(* Logix 5000 project; controller MV vendor 1 type 14 code 217 rev 31.11; software revision 31.00; part 31 of 53 *)
(* tags used below, declared in another part *)
   Alarm_Reset : BOOL;
   CWD : CHECKWORD_FLAGS;
   Default_Check_Time : DINT;
   Item_Faults_Are_Latched : BOOL;
   Item_Simulation_Flag : BOOL;
   MC_CD_T1 : PlantItem;   // CD_T1
   MC_CD_T1_ALARM : ALARM_DIGITAL;
   MC_CD_T1_C : ALIAS FOR RIO_Rack_2:7:I.Data.23;
   MC_CD_T1_DR : ALIAS FOR RIO_Rack_2:8:O.Data.11;
   MC_CD_T1_O : ALIAS FOR RIO_Rack_2:7:I.Data.19;
   MC_CD_T2 : PlantItem;   // CD_T2
   MC_CD_T2_ALARM : ALARM_DIGITAL;
   MC_CD_T2_C : ALIAS FOR RIO_Rack_2:7:I.Data.28;
   MC_CD_T2_DR : ALIAS FOR RIO_Rack_2:8:O.Data.12;
   MC_CD_T2_O : ALIAS FOR RIO_Rack_2:7:I.Data.24;
   MC_CH2_DR1 : PlantItem;   // CH2_DR1
   MC_CH2_DR1_ALARM : ALARM_DIGITAL;
   MC_CH2_DR1_C : ALIAS FOR RIO_Rack_2:7:I.Data.6;
   MC_CH2_DR1_DR : ALIAS FOR RIO_Rack_2:8:O.Data.2;
   MC_CH2_DR1_O : ALIAS FOR RIO_Rack_2:7:I.Data.2;
   MC_CH2_DR2 : PlantItem;   // CH2_DR2
   MC_CH2_DR2_ALARM : ALARM_DIGITAL;
   MC_CH2_DR2_C : ALIAS FOR RIO_Rack_2:7:I.Data.7;
   MC_CH2_DR2_DR : ALIAS FOR RIO_Rack_2:8:O.Data.3;
   MC_CH2_DR2_O : ALIAS FOR RIO_Rack_2:7:I.Data.3;
   MC_CH2_DRAIN : PlantItem;   // CH2_DRAIN
   MC_CH2_DRAIN_ALARM : ALARM_DIGITAL;
   MC_CH2_DRAIN_C : ALIAS FOR RIO_Rack_2:7:I.Data.4;
   MC_CH2_DRAIN_DR : ALIAS FOR RIO_Rack_2:8:O.Data.0;
   MC_CH2_DRAIN_O : ALIAS FOR RIO_Rack_2:7:I.Data.0;
   MC_CH2_DT1 : PlantItem;   // CH2_DT1
   MC_CH2_DT1_ALARM : ALARM_DIGITAL;
   MC_CH2_DT1_C : ALIAS FOR RIO_Rack_2:7:I.Data.12;
   MC_CH2_DT1_DR : ALIAS FOR RIO_Rack_2:8:O.Data.4;
   MC_CH2_DT1_O : ALIAS FOR RIO_Rack_2:7:I.Data.8;
   MC_CH2_DT2 : PlantItem;   // CH2_DT2
   MC_CH2_DT2_ALARM : ALARM_DIGITAL;
   MC_CH2_DT2_C : ALIAS FOR RIO_Rack_2:7:I.Data.13;
   MC_CH2_DT2_DR : ALIAS FOR RIO_Rack_2:8:O.Data.5;
   MC_CH2_DT2_O : ALIAS FOR RIO_Rack_2:7:I.Data.9;
   MC_CH2_LF1 : PlantItem;   // CH2_LF1
   MC_CH2_LF1_ALARM : ALARM_DIGITAL;
   MC_CH2_LF1_C : ALIAS FOR RIO_Rack_2:7:I.Data.15;
   MC_CH2_LF1_DR : ALIAS FOR RIO_Rack_2:8:O.Data.7;
   MC_CH2_LF1_O : ALIAS FOR RIO_Rack_2:7:I.Data.11;
   MC_CH2_PR1 : PlantItem;   // CH2_PR1
   MC_CH2_PR1_ALARM : ALARM_DIGITAL;
   MC_CH2_PR1_C : ALIAS FOR RIO_Rack_2:7:I.Data.14;
   MC_CH2_PR1_DR : ALIAS FOR RIO_Rack_2:8:O.Data.6;
   MC_CH2_PR1_O : ALIAS FOR RIO_Rack_2:7:I.Data.10;
   MC_CH2_R6R : PlantItem;   // CH2_R6R
   MC_CH2_R6R_ALARM : ALARM_DIGITAL;
   MC_CH2_R6R_C : ALIAS FOR RIO_Rack_2:6:I.Data.31;
   MC_CH2_R6R_DR : ALIAS FOR RIO_Rack_2:5:O.Data.31;
   MC_CH2_R6R_O : ALIAS FOR RIO_Rack_2:6:I.Data.27;
   MC_CH2_RR : PlantItem;   // CH2_RR
   MC_CH2_RR_ALARM : ALARM_DIGITAL;
   MC_CH2_RR_C : ALIAS FOR RIO_Rack_2:7:I.Data.5;
   MC_CH2_RR_DR : ALIAS FOR RIO_Rack_2:8:O.Data.1;
   MC_CH2_RR_O : ALIAS FOR RIO_Rack_2:7:I.Data.1;
   MC_FL_D1 : PlantItem;   // FL_D1
   MC_FL_D1_ALARM : ALARM_DIGITAL;
   MC_FL_D1_C : ALIAS FOR RIO_Rack_2:7:I.Data.21;
   MC_FL_D1_DR : ALIAS FOR RIO_Rack_2:8:O.Data.9;
   MC_FL_D1_O : ALIAS FOR RIO_Rack_2:7:I.Data.17;
   MC_FL_D2 : PlantItem;   // FL_D2
   MC_FL_D2_ALARM : ALARM_DIGITAL;
   MC_FL_D2_C : ALIAS FOR RIO_Rack_2:7:I.Data.22;
   MC_FL_D2_DR : ALIAS FOR RIO_Rack_2:8:O.Data.10;
   MC_FL_D2_O : ALIAS FOR RIO_Rack_2:7:I.Data.18;
   MC_FL_PR : PlantItem;   // FL_PR
   MC_FL_PR_ALARM : ALARM_DIGITAL;
   MC_FL_PR_C : ALIAS FOR RIO_Rack_2:7:I.Data.20;
   MC_FL_PR_DR : ALIAS FOR RIO_Rack_2:8:O.Data.8;
   MC_FL_PR_O : ALIAS FOR RIO_Rack_2:7:I.Data.16;
   MC_R3S_DR : PlantItem;   // R3S_DR
   MC_R3S_DR_ALARM : ALARM_DIGITAL;
   MC_R3S_DR_C : ALIAS FOR RIO_Rack_2:9:I.Data.15;
   MC_R3S_DR_DR : ALIAS FOR RIO_Rack_2:8:O.Data.23;
   MC_R3S_DR_O : ALIAS FOR RIO_Rack_2:9:I.Data.11;
   MC_R3V1 : PlantItem;   // R3V1
   MC_R3V1_ALARM : ALARM_DIGITAL;
   MC_R3V1_C : ALIAS FOR RIO_Rack_2:9:I.Data.12;
   MC_R3V1_DR : ALIAS FOR RIO_Rack_2:8:O.Data.20;
   MC_R3V1_O : ALIAS FOR RIO_Rack_2:9:I.Data.8;
   MC_R3V2 : PlantItem;   // R3V2
   MC_R3V2_ALARM : ALARM_DIGITAL;
   MC_R3V2_C : ALIAS FOR RIO_Rack_2:9:I.Data.13;
   MC_R3V2_DR : ALIAS FOR RIO_Rack_2:8:O.Data.21;
   MC_R3V2_O : ALIAS FOR RIO_Rack_2:9:I.Data.9;
   MC_SPV1 : PlantItem;   // SPV1
   MC_SPV1_ALARM : ALARM_DIGITAL;
   MC_SPV1_C : ALIAS FOR RIO_Rack_2:7:I.Data.31;
   MC_SPV1_DR : ALIAS FOR RIO_Rack_2:8:O.Data.15;
   MC_SPV1_O : ALIAS FOR RIO_Rack_2:7:I.Data.27;
   MC_SPV2 : PlantItem;   // SPV2
   MC_SPV2_ALARM : ALARM_DIGITAL;
   MC_SPV2_C : ALIAS FOR RIO_Rack_2:9:I.Data.4;
   MC_SPV2_DR : ALIAS FOR RIO_Rack_2:8:O.Data.16;
   MC_SPV2_O : ALIAS FOR RIO_Rack_2:9:I.Data.0;
   MC_SPV3 : PlantItem;   // SPV3
   MC_SPV3_ALARM : ALARM_DIGITAL;
   MC_SPV3_C : ALIAS FOR RIO_Rack_2:9:I.Data.5;
   MC_SPV3_DR : ALIAS FOR RIO_Rack_2:8:O.Data.17;
   MC_SPV3_O : ALIAS FOR RIO_Rack_2:9:I.Data.1;
   MC_SPV4 : PlantItem;   // SPV4
   MC_SPV4_ALARM : ALARM_DIGITAL;
   MC_SPV4_C : ALIAS FOR RIO_Rack_2:9:I.Data.6;
   MC_SPV4_DR : ALIAS FOR RIO_Rack_2:8:O.Data.18;
   MC_SPV4_O : ALIAS FOR RIO_Rack_2:9:I.Data.2;
   MC_SPV5 : PlantItem;   // SPV5
   MC_SPV5_ALARM : ALARM_DIGITAL;
   MC_SPV5_C : ALIAS FOR RIO_Rack_2:9:I.Data.7;
   MC_SPV5_DR : ALIAS FOR RIO_Rack_2:8:O.Data.19;
   MC_SPV5_O : ALIAS FOR RIO_Rack_2:9:I.Data.3;
   MC_SV1 : PlantItem;   // SV1
   MC_SV1_ALARM : ALARM_DIGITAL;
   MC_SV1_C : ALIAS FOR RIO_Rack_2:7:I.Data.29;
   MC_SV1_DR : ALIAS FOR RIO_Rack_2:8:O.Data.13;
   MC_SV1_O : ALIAS FOR RIO_Rack_2:7:I.Data.25;
   MC_SV2 : PlantItem;   // SV2
   MC_SV2_ALARM : ALARM_DIGITAL;
   MC_SV2_C : ALIAS FOR RIO_Rack_2:7:I.Data.30;
   MC_SV2_DR : ALIAS FOR RIO_Rack_2:8:O.Data.14;
   MC_SV2_O : ALIAS FOR RIO_Rack_2:7:I.Data.26;
   One_Second_One_Scan : ALIAS FOR One_Second_1_scan;
(* MC_Common, continued *)

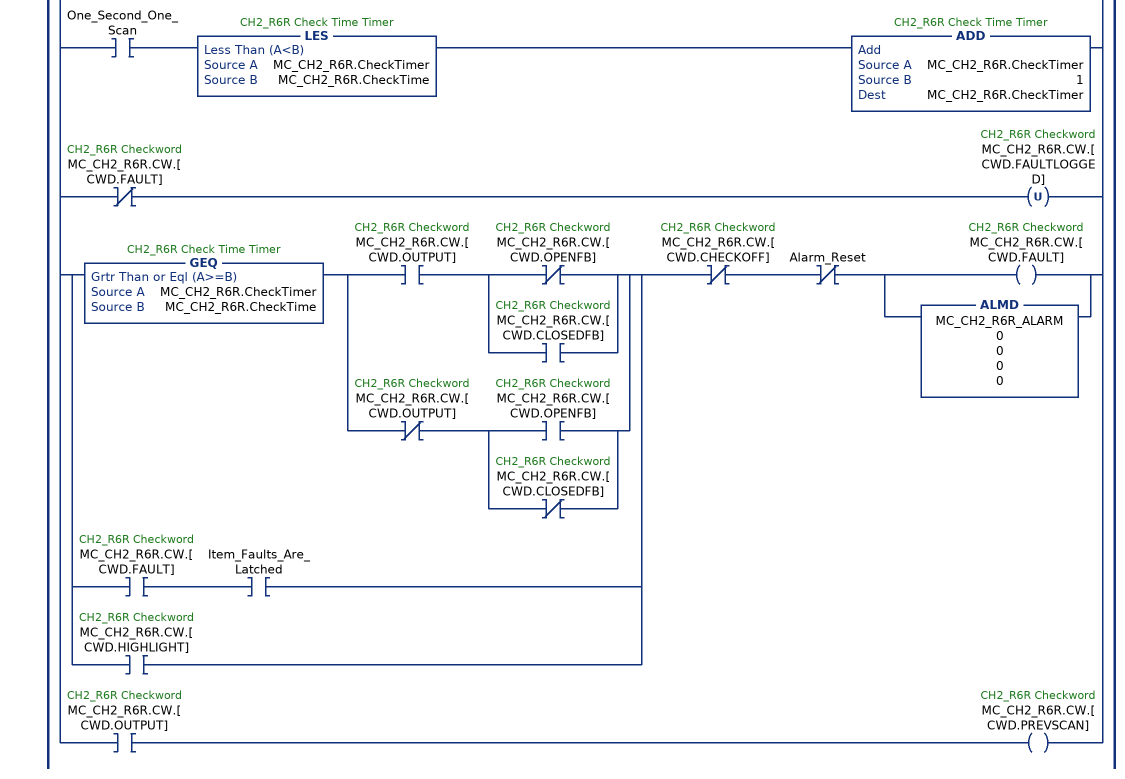
   [picture p660: MC_Common/MC_Valves rungs 31-31]
   31: [NEQ(MC_CH2_R6R.DriveBits,0) OTE(MC_CH2_R6R.CW.[CWD.AUTODRV]) ,[XIC(MC_CH2_R6R.CW.[CWD.AUTODRV]) XIO(MC_CH2_R6R.CW.[CWD.MANUAL]) ,XIC(MC_CH2_R6R.CW.[CWD.MANDRV]) XIC(MC_CH2_R6R.CW.[CWD.MANUAL]) ] OTE(MC_CH2_R6R.CW.[CWD.OUTPUT]) ,XIC(MC_CH2_R6R.CW.[CWD.OUTPUT]) OTE(MC_CH2_R6R_DR) ,XIC(S:FS) [OTU(MC_CH2_R6R.CW.[CWD.MANUAL]) ,LEQ(MC_CH2_R6R.CheckTime,0) MOV(Default_Check_Time,MC_CH2_R6R.CheckTime) ] ,[[XIC(MC_CH2_R6R_O) XIO(Item_Simulation_Flag) ,XIC(Item_Simulation_Flag) XIC(MC_CH2_R6R.CW.[CWD.OUTPUT]) XIO(MC_CH2_R6R.CW.[CWD.SIMFAIL]) ] OTE(MC_CH2_R6R.CW.[CWD.OPENFB]) ,[XIC(MC_CH2_R6R_C) XIO(Item_Simulation_Flag) ,XIC(Item_Simulation_Flag) XIO(MC_CH2_R6R.CW.[CWD.OUTPUT]) XIO(MC_CH2_R6R.CW.[CWD.SIMFAIL]) ] OTE(MC_CH2_R6R.CW.[CWD.CLOSEDFB]) ] ,[XIC(MC_CH2_R6R.CW.[CWD.OUTPUT]) XIO(MC_CH2_R6R.CW.[CWD.PREVSCAN]) ,XIO(MC_CH2_R6R.CW.[CWD.OUTPUT]) XIC(MC_CH2_R6R.CW.[CWD.PREVSCAN]) ] CLR(MC_CH2_R6R.CheckTimer) ,XIC(One_Second_One_Scan) LES(MC_CH2_R6R.CheckTimer,MC_CH2_R6R.CheckTime) ADD(MC_CH2_R6R.CheckTimer,1,MC_CH2_R6R.CheckTimer) ,XIO(MC_CH2_R6R.CW.[CWD.FAULT]) OTU(MC_CH2_R6R.CW.[CWD.FAULTLOGGED]) ,[GEQ(MC_CH2_R6R.CheckTimer,MC_CH2_R6R.CheckTime) [XIC(MC_CH2_R6R.CW.[CWD.OUTPUT]) [XIO(MC_CH2_R6R.CW.[CWD.OPENFB]) ,XIC(MC_CH2_R6R.CW.[CWD.CLOSEDFB]) ] ,XIO(MC_CH2_R6R.CW.[CWD.OUTPUT]) [XIC(MC_CH2_R6R.CW.[CWD.OPENFB]) ,XIO(MC_CH2_R6R.CW.[CWD.CLOSEDFB]) ] ] ,XIC(MC_CH2_R6R.CW.[CWD.FAULT]) XIC(Item_Faults_Are_Latched) ,XIC(MC_CH2_R6R.CW.[CWD.HIGHLIGHT]) ] XIO(MC_CH2_R6R.CW.[CWD.CHECKOFF]) XIO(Alarm_Reset) [OTE(MC_CH2_R6R.CW.[CWD.FAULT]) ,ALMD(MC_CH2_R6R_ALARM,0,0,0,0) ] ,XIC(MC_CH2_R6R.CW.[CWD.OUTPUT]) OTE(MC_CH2_R6R.CW.[CWD.PREVSCAN]) ];
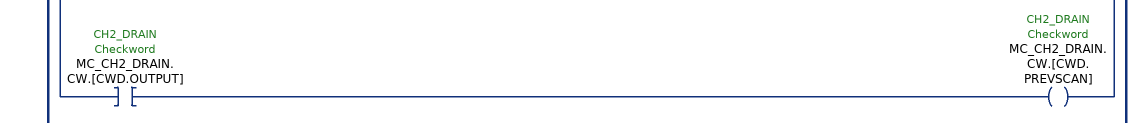
   32: [NEQ(MC_CH2_DRAIN.DriveBits,0) OTE(MC_CH2_DRAIN.CW.[CWD.AUTODRV]) ,[XIC(MC_CH2_DRAIN.CW.[CWD.AUTODRV]) XIO(MC_CH2_DRAIN.CW.[CWD.MANUAL]) ,XIC(MC_CH2_DRAIN.CW.[CWD.MANDRV]) XIC(MC_CH2_DRAIN.CW.[CWD.MANUAL]) ] OTE(MC_CH2_DRAIN.CW.[CWD.OUTPUT]) ,XIC(MC_CH2_DRAIN.CW.[CWD.OUTPUT]) OTE(MC_CH2_DRAIN_DR) ,XIC(S:FS) [OTU(MC_CH2_DRAIN.CW.[CWD.MANUAL]) ,LEQ(MC_CH2_DRAIN.CheckTime,0) MOV(Default_Check_Time,MC_CH2_DRAIN.CheckTime) ] ,[[XIC(MC_CH2_DRAIN_O) XIO(Item_Simulation_Flag) ,XIC(Item_Simulation_Flag) XIC(MC_CH2_DRAIN.CW.[CWD.OUTPUT]) XIO(MC_CH2_DRAIN.CW.[CWD.SIMFAIL]) ] OTE(MC_CH2_DRAIN.CW.[CWD.OPENFB]) ,[XIC(MC_CH2_DRAIN_C) XIO(Item_Simulation_Flag) ,XIC(Item_Simulation_Flag) XIO(MC_CH2_DRAIN.CW.[CWD.OUTPUT]) XIO(MC_CH2_DRAIN.CW.[CWD.SIMFAIL]) ] OTE(MC_CH2_DRAIN.CW.[CWD.CLOSEDFB]) ] ,[XIC(MC_CH2_DRAIN.CW.[CWD.OUTPUT]) XIO(MC_CH2_DRAIN.CW.[CWD.PREVSCAN]) ,XIO(MC_CH2_DRAIN.CW.[CWD.OUTPUT]) XIC(MC_CH2_DRAIN.CW.[CWD.PREVSCAN]) ] CLR(MC_CH2_DRAIN.CheckTimer) ,XIC(One_Second_One_Scan) LES(MC_CH2_DRAIN.CheckTimer,MC_CH2_DRAIN.CheckTime) ADD(MC_CH2_DRAIN.CheckTimer,1,MC_CH2_DRAIN.CheckTimer) ,XIO(MC_CH2_DRAIN.CW.[CWD.FAULT]) OTU(MC_CH2_DRAIN.CW.[CWD.FAULTLOGGED]) ,[GEQ(MC_CH2_DRAIN.CheckTimer,MC_CH2_DRAIN.CheckTime) [XIC(MC_CH2_DRAIN.CW.[CWD.OUTPUT]) [XIO(MC_CH2_DRAIN.CW.[CWD.OPENFB]) ,XIC(MC_CH2_DRAIN.CW.[CWD.CLOSEDFB]) ] ,XIO(MC_CH2_DRAIN.CW.[CWD.OUTPUT]) [XIC(MC_CH2_DRAIN.CW.[CWD.OPENFB]) ,XIO(MC_CH2_DRAIN.CW.[CWD.CLOSEDFB]) ] ] ,XIC(MC_CH2_DRAIN.CW.[CWD.FAULT]) XIC(Item_Faults_Are_Latched) ,XIC(MC_CH2_DRAIN.CW.[CWD.HIGHLIGHT]) ] XIO(MC_CH2_DRAIN.CW.[CWD.CHECKOFF]) XIO(Alarm_Reset) [OTE(MC_CH2_DRAIN.CW.[CWD.FAULT]) ,ALMD(MC_CH2_DRAIN_ALARM,0,0,0,0) ] ,XIC(MC_CH2_DRAIN.CW.[CWD.OUTPUT]) OTE(MC_CH2_DRAIN.CW.[CWD.PREVSCAN]) ];
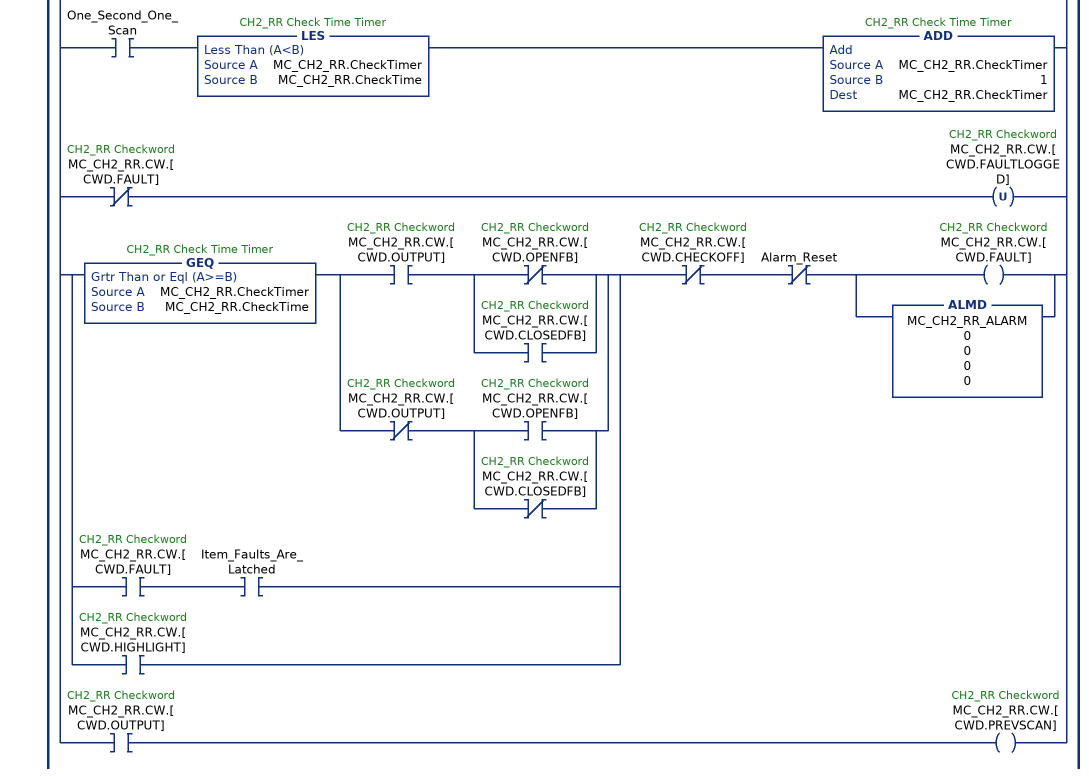
   33: [NEQ(MC_CH2_RR.DriveBits,0) OTE(MC_CH2_RR.CW.[CWD.AUTODRV]) ,[XIC(MC_CH2_RR.CW.[CWD.AUTODRV]) XIO(MC_CH2_RR.CW.[CWD.MANUAL]) ,XIC(MC_CH2_RR.CW.[CWD.MANDRV]) XIC(MC_CH2_RR.CW.[CWD.MANUAL]) ] OTE(MC_CH2_RR.CW.[CWD.OUTPUT]) ,XIC(MC_CH2_RR.CW.[CWD.OUTPUT]) OTE(MC_CH2_RR_DR) ,XIC(S:FS) [OTU(MC_CH2_RR.CW.[CWD.MANUAL]) ,LEQ(MC_CH2_RR.CheckTime,0) MOV(Default_Check_Time,MC_CH2_RR.CheckTime) ] ,[[XIC(MC_CH2_RR_O) XIO(Item_Simulation_Flag) ,XIC(Item_Simulation_Flag) XIC(MC_CH2_RR.CW.[CWD.OUTPUT]) XIO(MC_CH2_RR.CW.[CWD.SIMFAIL]) ] OTE(MC_CH2_RR.CW.[CWD.OPENFB]) ,[XIC(MC_CH2_RR_C) XIO(Item_Simulation_Flag) ,XIC(Item_Simulation_Flag) XIO(MC_CH2_RR.CW.[CWD.OUTPUT]) XIO(MC_CH2_RR.CW.[CWD.SIMFAIL]) ] OTE(MC_CH2_RR.CW.[CWD.CLOSEDFB]) ] ,[XIC(MC_CH2_RR.CW.[CWD.OUTPUT]) XIO(MC_CH2_RR.CW.[CWD.PREVSCAN]) ,XIO(MC_CH2_RR.CW.[CWD.OUTPUT]) XIC(MC_CH2_RR.CW.[CWD.PREVSCAN]) ] CLR(MC_CH2_RR.CheckTimer) ,XIC(One_Second_One_Scan) LES(MC_CH2_RR.CheckTimer,MC_CH2_RR.CheckTime) ADD(MC_CH2_RR.CheckTimer,1,MC_CH2_RR.CheckTimer) ,XIO(MC_CH2_RR.CW.[CWD.FAULT]) OTU(MC_CH2_RR.CW.[CWD.FAULTLOGGED]) ,[GEQ(MC_CH2_RR.CheckTimer,MC_CH2_RR.CheckTime) [XIC(MC_CH2_RR.CW.[CWD.OUTPUT]) [XIO(MC_CH2_RR.CW.[CWD.OPENFB]) ,XIC(MC_CH2_RR.CW.[CWD.CLOSEDFB]) ] ,XIO(MC_CH2_RR.CW.[CWD.OUTPUT]) [XIC(MC_CH2_RR.CW.[CWD.OPENFB]) ,XIO(MC_CH2_RR.CW.[CWD.CLOSEDFB]) ] ] ,XIC(MC_CH2_RR.CW.[CWD.FAULT]) XIC(Item_Faults_Are_Latched) ,XIC(MC_CH2_RR.CW.[CWD.HIGHLIGHT]) ] XIO(MC_CH2_RR.CW.[CWD.CHECKOFF]) XIO(Alarm_Reset) [OTE(MC_CH2_RR.CW.[CWD.FAULT]) ,ALMD(MC_CH2_RR_ALARM,0,0,0,0) ] ,XIC(MC_CH2_RR.CW.[CWD.OUTPUT]) OTE(MC_CH2_RR.CW.[CWD.PREVSCAN]) ];
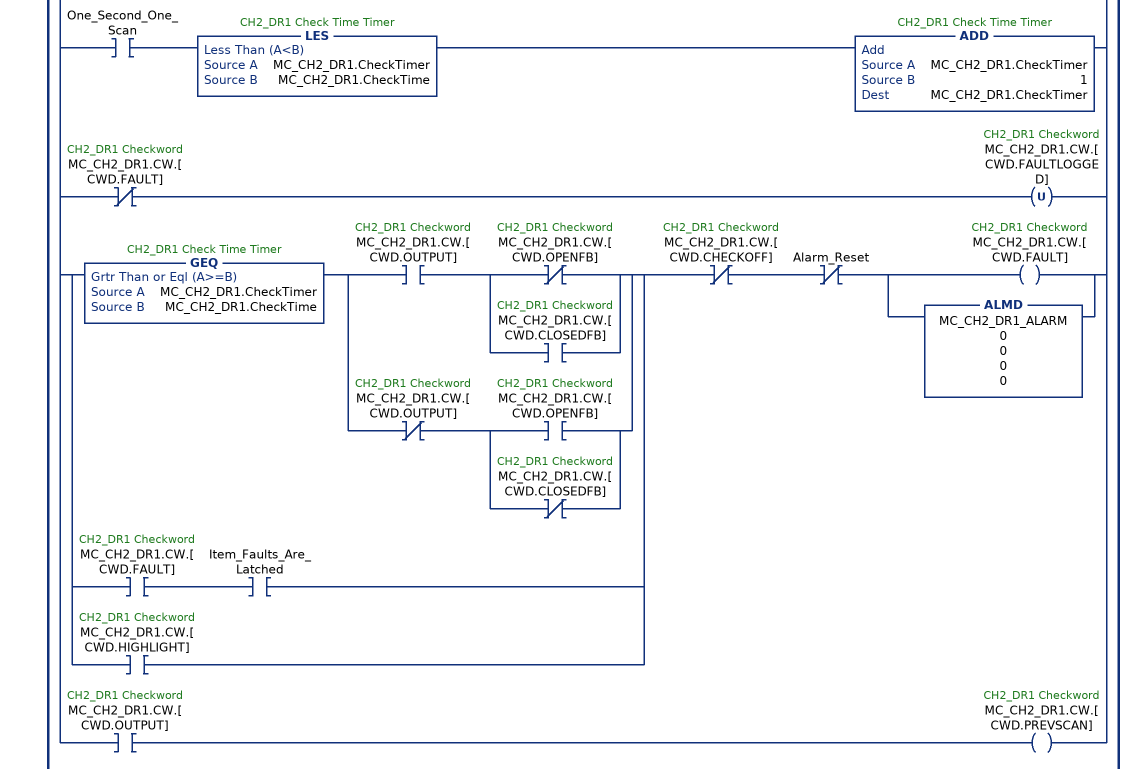
   34: [NEQ(MC_CH2_DR1.DriveBits,0) OTE(MC_CH2_DR1.CW.[CWD.AUTODRV]) ,[XIC(MC_CH2_DR1.CW.[CWD.AUTODRV]) XIO(MC_CH2_DR1.CW.[CWD.MANUAL]) ,XIC(MC_CH2_DR1.CW.[CWD.MANDRV]) XIC(MC_CH2_DR1.CW.[CWD.MANUAL]) ] OTE(MC_CH2_DR1.CW.[CWD.OUTPUT]) ,XIC(MC_CH2_DR1.CW.[CWD.OUTPUT]) OTE(MC_CH2_DR1_DR) ,XIC(S:FS) [OTU(MC_CH2_DR1.CW.[CWD.MANUAL]) ,LEQ(MC_CH2_DR1.CheckTime,0) MOV(Default_Check_Time,MC_CH2_DR1.CheckTime) ] ,[[XIC(MC_CH2_DR1_O) XIO(Item_Simulation_Flag) ,XIC(Item_Simulation_Flag) XIC(MC_CH2_DR1.CW.[CWD.OUTPUT]) XIO(MC_CH2_DR1.CW.[CWD.SIMFAIL]) ] OTE(MC_CH2_DR1.CW.[CWD.OPENFB]) ,[XIC(MC_CH2_DR1_C) XIO(Item_Simulation_Flag) ,XIC(Item_Simulation_Flag) XIO(MC_CH2_DR1.CW.[CWD.OUTPUT]) XIO(MC_CH2_DR1.CW.[CWD.SIMFAIL]) ] OTE(MC_CH2_DR1.CW.[CWD.CLOSEDFB]) ] ,[XIC(MC_CH2_DR1.CW.[CWD.OUTPUT]) XIO(MC_CH2_DR1.CW.[CWD.PREVSCAN]) ,XIO(MC_CH2_DR1.CW.[CWD.OUTPUT]) XIC(MC_CH2_DR1.CW.[CWD.PREVSCAN]) ] CLR(MC_CH2_DR1.CheckTimer) ,XIC(One_Second_One_Scan) LES(MC_CH2_DR1.CheckTimer,MC_CH2_DR1.CheckTime) ADD(MC_CH2_DR1.CheckTimer,1,MC_CH2_DR1.CheckTimer) ,XIO(MC_CH2_DR1.CW.[CWD.FAULT]) OTU(MC_CH2_DR1.CW.[CWD.FAULTLOGGED]) ,[GEQ(MC_CH2_DR1.CheckTimer,MC_CH2_DR1.CheckTime) [XIC(MC_CH2_DR1.CW.[CWD.OUTPUT]) [XIO(MC_CH2_DR1.CW.[CWD.OPENFB]) ,XIC(MC_CH2_DR1.CW.[CWD.CLOSEDFB]) ] ,XIO(MC_CH2_DR1.CW.[CWD.OUTPUT]) [XIC(MC_CH2_DR1.CW.[CWD.OPENFB]) ,XIO(MC_CH2_DR1.CW.[CWD.CLOSEDFB]) ] ] ,XIC(MC_CH2_DR1.CW.[CWD.FAULT]) XIC(Item_Faults_Are_Latched) ,XIC(MC_CH2_DR1.CW.[CWD.HIGHLIGHT]) ] XIO(MC_CH2_DR1.CW.[CWD.CHECKOFF]) XIO(Alarm_Reset) [OTE(MC_CH2_DR1.CW.[CWD.FAULT]) ,ALMD(MC_CH2_DR1_ALARM,0,0,0,0) ] ,XIC(MC_CH2_DR1.CW.[CWD.OUTPUT]) OTE(MC_CH2_DR1.CW.[CWD.PREVSCAN]) ];
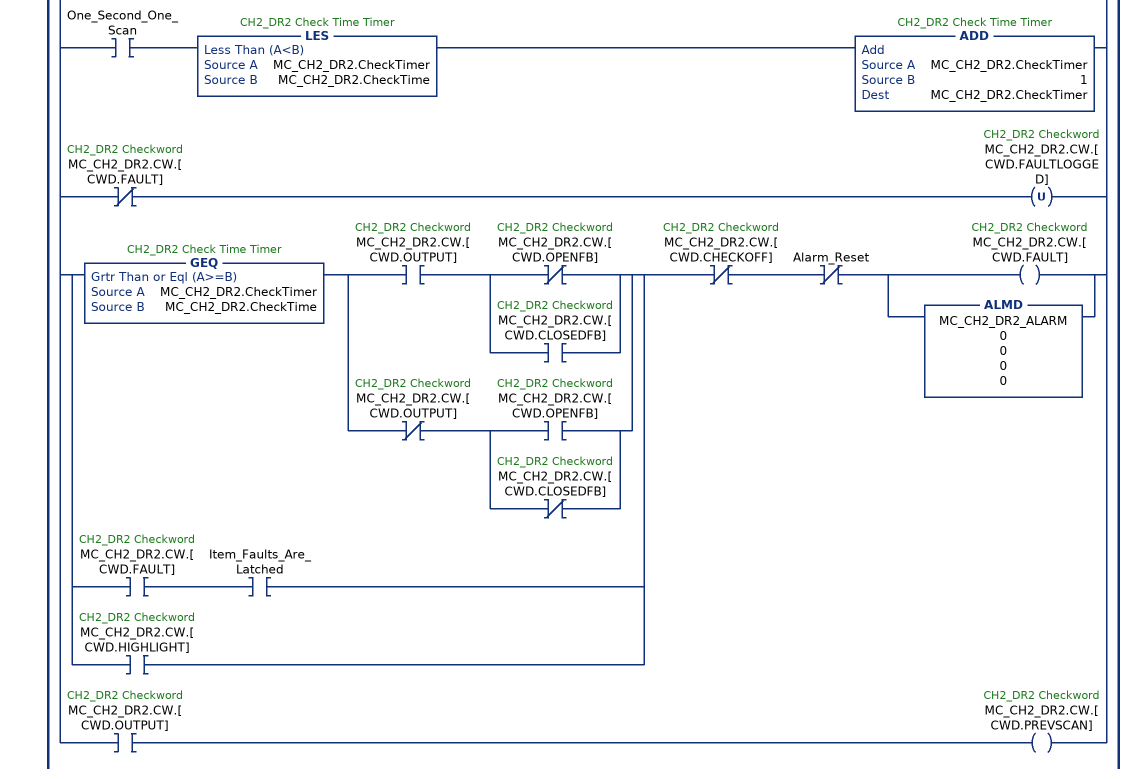
   35: [NEQ(MC_CH2_DR2.DriveBits,0) OTE(MC_CH2_DR2.CW.[CWD.AUTODRV]) ,[XIC(MC_CH2_DR2.CW.[CWD.AUTODRV]) XIO(MC_CH2_DR2.CW.[CWD.MANUAL]) ,XIC(MC_CH2_DR2.CW.[CWD.MANDRV]) XIC(MC_CH2_DR2.CW.[CWD.MANUAL]) ] OTE(MC_CH2_DR2.CW.[CWD.OUTPUT]) ,XIC(MC_CH2_DR2.CW.[CWD.OUTPUT]) OTE(MC_CH2_DR2_DR) ,XIC(S:FS) [OTU(MC_CH2_DR2.CW.[CWD.MANUAL]) ,LEQ(MC_CH2_DR2.CheckTime,0) MOV(Default_Check_Time,MC_CH2_DR2.CheckTime) ] ,[[XIC(MC_CH2_DR2_O) XIO(Item_Simulation_Flag) ,XIC(Item_Simulation_Flag) XIC(MC_CH2_DR2.CW.[CWD.OUTPUT]) XIO(MC_CH2_DR2.CW.[CWD.SIMFAIL]) ] OTE(MC_CH2_DR2.CW.[CWD.OPENFB]) ,[XIC(MC_CH2_DR2_C) XIO(Item_Simulation_Flag) ,XIC(Item_Simulation_Flag) XIO(MC_CH2_DR2.CW.[CWD.OUTPUT]) XIO(MC_CH2_DR2.CW.[CWD.SIMFAIL]) ] OTE(MC_CH2_DR2.CW.[CWD.CLOSEDFB]) ] ,[XIC(MC_CH2_DR2.CW.[CWD.OUTPUT]) XIO(MC_CH2_DR2.CW.[CWD.PREVSCAN]) ,XIO(MC_CH2_DR2.CW.[CWD.OUTPUT]) XIC(MC_CH2_DR2.CW.[CWD.PREVSCAN]) ] CLR(MC_CH2_DR2.CheckTimer) ,XIC(One_Second_One_Scan) LES(MC_CH2_DR2.CheckTimer,MC_CH2_DR2.CheckTime) ADD(MC_CH2_DR2.CheckTimer,1,MC_CH2_DR2.CheckTimer) ,XIO(MC_CH2_DR2.CW.[CWD.FAULT]) OTU(MC_CH2_DR2.CW.[CWD.FAULTLOGGED]) ,[GEQ(MC_CH2_DR2.CheckTimer,MC_CH2_DR2.CheckTime) [XIC(MC_CH2_DR2.CW.[CWD.OUTPUT]) [XIO(MC_CH2_DR2.CW.[CWD.OPENFB]) ,XIC(MC_CH2_DR2.CW.[CWD.CLOSEDFB]) ] ,XIO(MC_CH2_DR2.CW.[CWD.OUTPUT]) [XIC(MC_CH2_DR2.CW.[CWD.OPENFB]) ,XIO(MC_CH2_DR2.CW.[CWD.CLOSEDFB]) ] ] ,XIC(MC_CH2_DR2.CW.[CWD.FAULT]) XIC(Item_Faults_Are_Latched) ,XIC(MC_CH2_DR2.CW.[CWD.HIGHLIGHT]) ] XIO(MC_CH2_DR2.CW.[CWD.CHECKOFF]) XIO(Alarm_Reset) [OTE(MC_CH2_DR2.CW.[CWD.FAULT]) ,ALMD(MC_CH2_DR2_ALARM,0,0,0,0) ] ,XIC(MC_CH2_DR2.CW.[CWD.OUTPUT]) OTE(MC_CH2_DR2.CW.[CWD.PREVSCAN]) ];
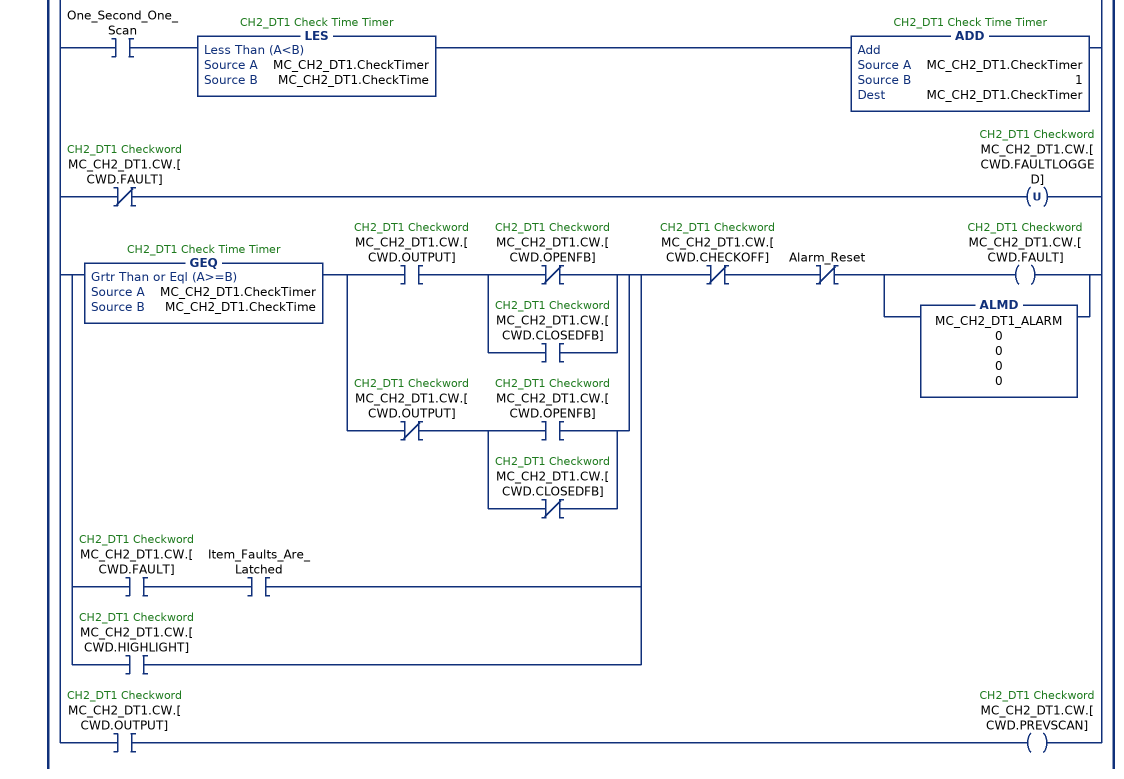
   36: [NEQ(MC_CH2_DT1.DriveBits,0) OTE(MC_CH2_DT1.CW.[CWD.AUTODRV]) ,[XIC(MC_CH2_DT1.CW.[CWD.AUTODRV]) XIO(MC_CH2_DT1.CW.[CWD.MANUAL]) ,XIC(MC_CH2_DT1.CW.[CWD.MANDRV]) XIC(MC_CH2_DT1.CW.[CWD.MANUAL]) ] OTE(MC_CH2_DT1.CW.[CWD.OUTPUT]) ,XIC(MC_CH2_DT1.CW.[CWD.OUTPUT]) OTE(MC_CH2_DT1_DR) ,XIC(S:FS) [OTU(MC_CH2_DT1.CW.[CWD.MANUAL]) ,LEQ(MC_CH2_DT1.CheckTime,0) MOV(Default_Check_Time,MC_CH2_DT1.CheckTime) ] ,[[XIC(MC_CH2_DT1_O) XIO(Item_Simulation_Flag) ,XIC(Item_Simulation_Flag) XIC(MC_CH2_DT1.CW.[CWD.OUTPUT]) XIO(MC_CH2_DT1.CW.[CWD.SIMFAIL]) ] OTE(MC_CH2_DT1.CW.[CWD.OPENFB]) ,[XIC(MC_CH2_DT1_C) XIO(Item_Simulation_Flag) ,XIC(Item_Simulation_Flag) XIO(MC_CH2_DT1.CW.[CWD.OUTPUT]) XIO(MC_CH2_DT1.CW.[CWD.SIMFAIL]) ] OTE(MC_CH2_DT1.CW.[CWD.CLOSEDFB]) ] ,[XIC(MC_CH2_DT1.CW.[CWD.OUTPUT]) XIO(MC_CH2_DT1.CW.[CWD.PREVSCAN]) ,XIO(MC_CH2_DT1.CW.[CWD.OUTPUT]) XIC(MC_CH2_DT1.CW.[CWD.PREVSCAN]) ] CLR(MC_CH2_DT1.CheckTimer) ,XIC(One_Second_One_Scan) LES(MC_CH2_DT1.CheckTimer,MC_CH2_DT1.CheckTime) ADD(MC_CH2_DT1.CheckTimer,1,MC_CH2_DT1.CheckTimer) ,XIO(MC_CH2_DT1.CW.[CWD.FAULT]) OTU(MC_CH2_DT1.CW.[CWD.FAULTLOGGED]) ,[GEQ(MC_CH2_DT1.CheckTimer,MC_CH2_DT1.CheckTime) [XIC(MC_CH2_DT1.CW.[CWD.OUTPUT]) [XIO(MC_CH2_DT1.CW.[CWD.OPENFB]) ,XIC(MC_CH2_DT1.CW.[CWD.CLOSEDFB]) ] ,XIO(MC_CH2_DT1.CW.[CWD.OUTPUT]) [XIC(MC_CH2_DT1.CW.[CWD.OPENFB]) ,XIO(MC_CH2_DT1.CW.[CWD.CLOSEDFB]) ] ] ,XIC(MC_CH2_DT1.CW.[CWD.FAULT]) XIC(Item_Faults_Are_Latched) ,XIC(MC_CH2_DT1.CW.[CWD.HIGHLIGHT]) ] XIO(MC_CH2_DT1.CW.[CWD.CHECKOFF]) XIO(Alarm_Reset) [OTE(MC_CH2_DT1.CW.[CWD.FAULT]) ,ALMD(MC_CH2_DT1_ALARM,0,0,0,0) ] ,XIC(MC_CH2_DT1.CW.[CWD.OUTPUT]) OTE(MC_CH2_DT1.CW.[CWD.PREVSCAN]) ];
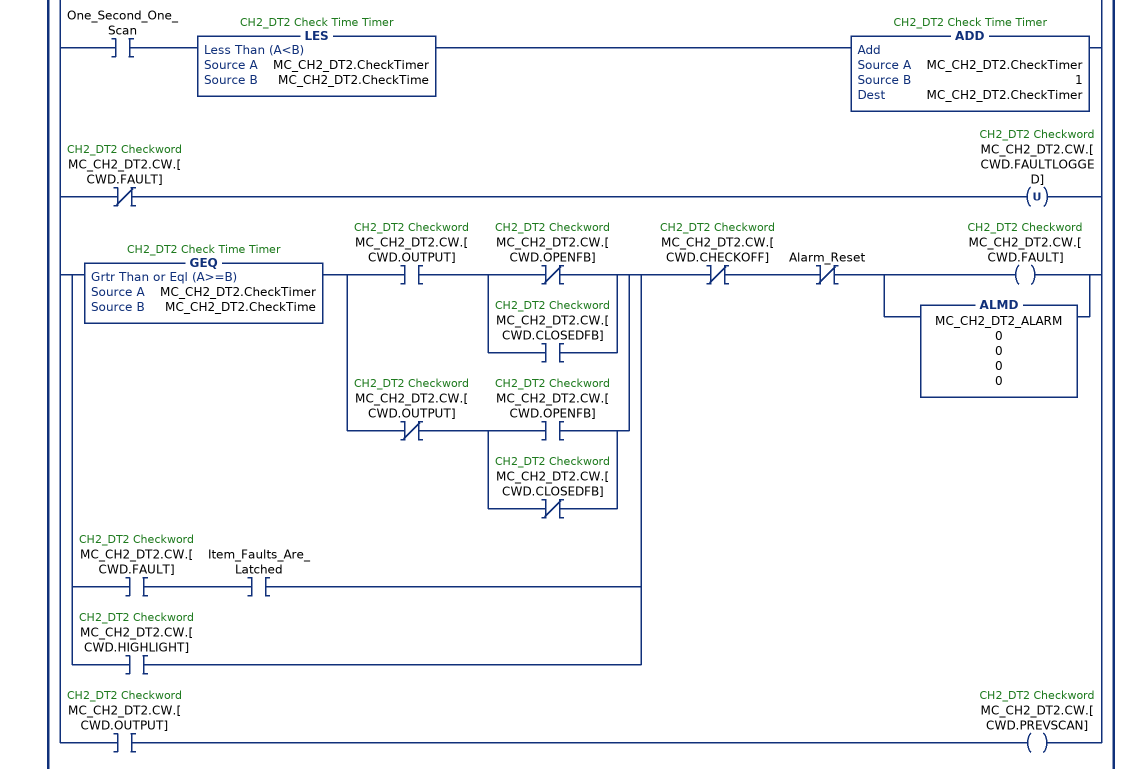
   37: [NEQ(MC_CH2_DT2.DriveBits,0) OTE(MC_CH2_DT2.CW.[CWD.AUTODRV]) ,[XIC(MC_CH2_DT2.CW.[CWD.AUTODRV]) XIO(MC_CH2_DT2.CW.[CWD.MANUAL]) ,XIC(MC_CH2_DT2.CW.[CWD.MANDRV]) XIC(MC_CH2_DT2.CW.[CWD.MANUAL]) ] OTE(MC_CH2_DT2.CW.[CWD.OUTPUT]) ,XIC(MC_CH2_DT2.CW.[CWD.OUTPUT]) OTE(MC_CH2_DT2_DR) ,XIC(S:FS) [OTU(MC_CH2_DT2.CW.[CWD.MANUAL]) ,LEQ(MC_CH2_DT2.CheckTime,0) MOV(Default_Check_Time,MC_CH2_DT2.CheckTime) ] ,[[XIC(MC_CH2_DT2_O) XIO(Item_Simulation_Flag) ,XIC(Item_Simulation_Flag) XIC(MC_CH2_DT2.CW.[CWD.OUTPUT]) XIO(MC_CH2_DT2.CW.[CWD.SIMFAIL]) ] OTE(MC_CH2_DT2.CW.[CWD.OPENFB]) ,[XIC(MC_CH2_DT2_C) XIO(Item_Simulation_Flag) ,XIC(Item_Simulation_Flag) XIO(MC_CH2_DT2.CW.[CWD.OUTPUT]) XIO(MC_CH2_DT2.CW.[CWD.SIMFAIL]) ] OTE(MC_CH2_DT2.CW.[CWD.CLOSEDFB]) ] ,[XIC(MC_CH2_DT2.CW.[CWD.OUTPUT]) XIO(MC_CH2_DT2.CW.[CWD.PREVSCAN]) ,XIO(MC_CH2_DT2.CW.[CWD.OUTPUT]) XIC(MC_CH2_DT2.CW.[CWD.PREVSCAN]) ] CLR(MC_CH2_DT2.CheckTimer) ,XIC(One_Second_One_Scan) LES(MC_CH2_DT2.CheckTimer,MC_CH2_DT2.CheckTime) ADD(MC_CH2_DT2.CheckTimer,1,MC_CH2_DT2.CheckTimer) ,XIO(MC_CH2_DT2.CW.[CWD.FAULT]) OTU(MC_CH2_DT2.CW.[CWD.FAULTLOGGED]) ,[GEQ(MC_CH2_DT2.CheckTimer,MC_CH2_DT2.CheckTime) [XIC(MC_CH2_DT2.CW.[CWD.OUTPUT]) [XIO(MC_CH2_DT2.CW.[CWD.OPENFB]) ,XIC(MC_CH2_DT2.CW.[CWD.CLOSEDFB]) ] ,XIO(MC_CH2_DT2.CW.[CWD.OUTPUT]) [XIC(MC_CH2_DT2.CW.[CWD.OPENFB]) ,XIO(MC_CH2_DT2.CW.[CWD.CLOSEDFB]) ] ] ,XIC(MC_CH2_DT2.CW.[CWD.FAULT]) XIC(Item_Faults_Are_Latched) ,XIC(MC_CH2_DT2.CW.[CWD.HIGHLIGHT]) ] XIO(MC_CH2_DT2.CW.[CWD.CHECKOFF]) XIO(Alarm_Reset) [OTE(MC_CH2_DT2.CW.[CWD.FAULT]) ,ALMD(MC_CH2_DT2_ALARM,0,0,0,0) ] ,XIC(MC_CH2_DT2.CW.[CWD.OUTPUT]) OTE(MC_CH2_DT2.CW.[CWD.PREVSCAN]) ];